   RUNG wire#powerrail
      Contact( "pH-2021_DB".Alarms.HighHigh )
   END_RUNG wire#w20
   RUNG wire#powerrail
      { S7_Templates := "SrcType := Time" } GE_Contact(in1 := "VFD-R201_DB".TIMEOUT.PT, in2 := T#8s)
   END_RUNG wire#w21
   RUNG wire#powerrail
      { S7_Templates := "SrcType := Time" } GE_Contact(in1 := "P-201A_DB".CF_Delay_TON.ET, in2 := T#8s)
   END_RUNG wire#w22
   RUNG wire#powerrail
      { S7_Templates := "SrcType := Time" } GE_Contact(in1 := "P-201B_DB".CF_Delay_TON.ET, in2 := T#8s)
   END_RUNG wire#w23
   RUNG wire#powerrail
      I_Contact( "T-101_Interlocks_DB".Out )
      P_Trig( "R-201_DB".OS.bit[1] )
   END_RUNG wire#w24
   // the same network as SCL:
   #_w1 := NOT "T-101_Interlocks_DB".Out AND NOT "R-201_DB".OS.bit[1];   // rising edge
   "R-201_DB".OS.bit[1] := NOT "T-101_Interlocks_DB".Out;
   "R-201_Interlocks_DB"(Interlock_1 := "LT-2011_DB".Alarms.HighHigh,   // "Interlocks"
                         Interlock_2 := "LSHH-2011_DB".Q,
                         Interlock_3 := "PT-201A_DB".Alarms.HighHigh,
                         Interlock_4 := "PT-201B_DB".Alarms.HighHigh,
                         Interlock_5 := "LT-2011_DB".Alarms.TransmitterFault,
                         Interlock_6 := "PT-201A_DB".Alarms.TransmitterFault,
                         Interlock_7 := "PT-201B_DB".Alarms.TransmitterFault,
                         Interlock_8 := "TT-2011_DB".Alarms.TransmitterFault,
                         Interlock_9 := "TT-2012_DB".Alarms.TransmitterFault,
                         Interlock_10 := "pH-2011_DB".Alarms.TransmitterFault,
                         Interlock_11 := "pH-2012_DB".Alarms.TransmitterFault,
                         Interlock_12 := "FT-2011_DB".Alarms.TransmitterFault,
                         Interlock_13 := "FT-2021_DB".Alarms.TransmitterFault,
                         Interlock_14 := "XV-2021_DB".Alarms."TO" OR "XV-2021_DB".Alarms.TC,
                         Interlock_15 := "XV-2013_DB".Alarms."TO" OR "XV-2013_DB".Alarms.TC,
                         Interlock_16 := "XV-1043_DB".Alarms."TO" OR "XV-1043_DB".Alarms.TC,
                         Interlock_17 := "XV-2011_DB".Alarms."TO" OR "XV-2011_DB".Alarms.TC,
                         Interlock_18 := "FT-1043_DB".Alarms.TransmitterFault,
                         Interlock_19 := "pH-2022_DB".Alarms.HighHigh,
                         Interlock_20 := "pH-2021_DB".Alarms.HighHigh,
                         Interlock_21 := "VFD-R201_DB".TIMEOUT.PT >= T#8s,
                         Interlock_22 := "P-201A_DB".CF_Delay_TON.ET >= T#8s,
                         Interlock_23 := "P-201B_DB".CF_Delay_TON.ET >= T#8s,
                         Interlock_25 := #_w1);
END_REGION

REGION Network 2: R-202 as Unit Interlocks
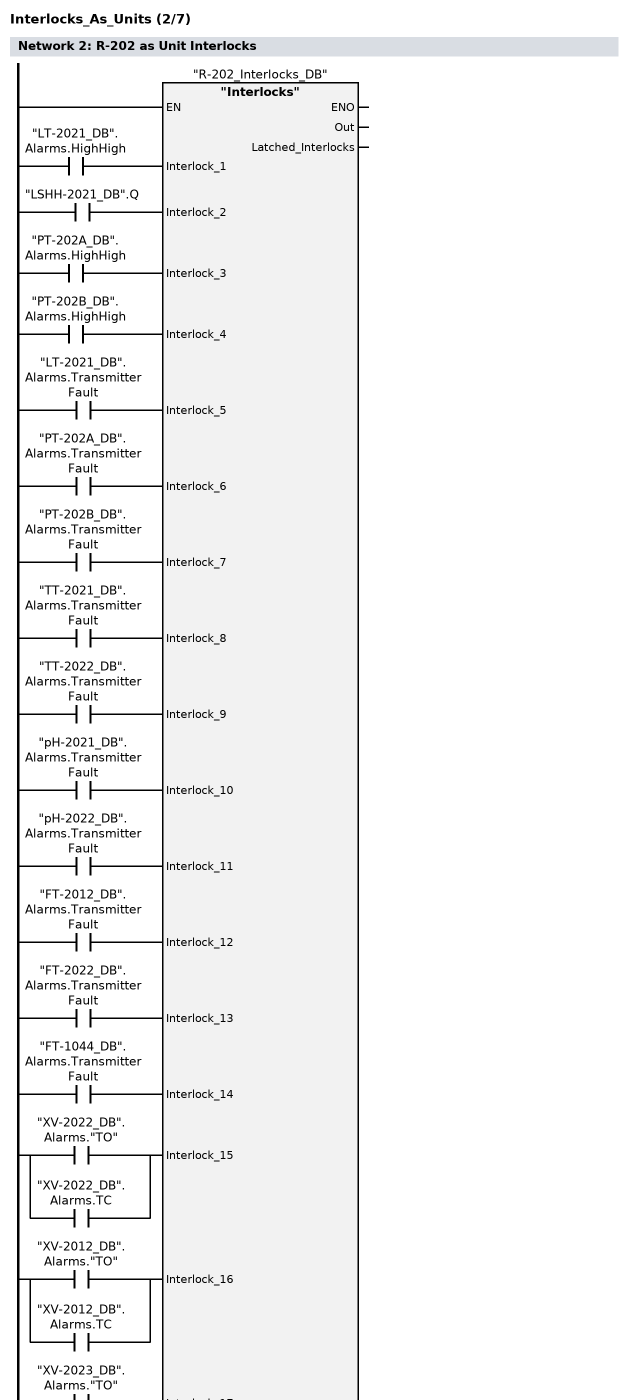
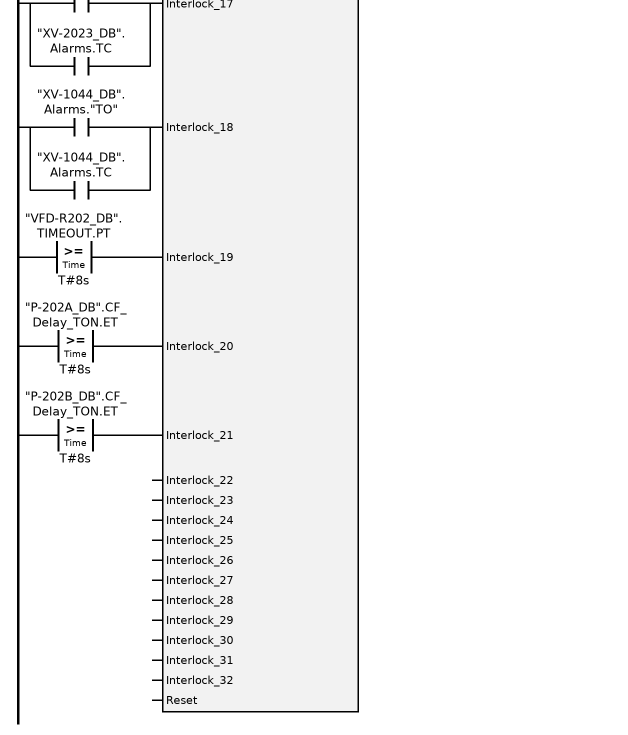
   RUNG wire#powerrail
      "R-202_Interlocks_DB"(Interlock_1 := wire#w1, Interlock_2 := wire#w2, Interlock_3 := wire#w3, Interlock_4 := wire#w4, Interlock_5 := wire#w5, Interlock_6 := wire#w6, Interlock_7 := wire#w7, Interlock_8 := wire#w8, Interlock_9 := wire#w9, Interlock_10 := wire#w10, Interlock_11 := wire#w11, Interlock_12 := wire#w12, Interlock_13 := wire#w13, Interlock_14 := wire#w14, Interlock_15 := wire#w15, Interlock_16 := wire#w16, Interlock_17 := wire#w17, Interlock_18 := wire#w18, Interlock_19 := wire#w19, Interlock_20 := wire#w20, Interlock_21 := wire#w21, Interlock_22 :=, Interlock_23 :=, Interlock_24 :=, Interlock_25 :=, Interlock_26 :=, Interlock_27 :=, Interlock_28 :=, Interlock_29 :=, Interlock_30 :=, Interlock_31 :=, Interlock_32 :=, Reset :=, Out =>, Latched_Interlocks =>)
   END_RUNG
   RUNG wire#powerrail
      Contact( "LT-2021_DB".Alarms.HighHigh )
   END_RUNG wire#w1
   RUNG wire#powerrail
      Contact( "LSHH-2021_DB".Q )
   END_RUNG wire#w2
   RUNG wire#powerrail
      Contact( "PT-202A_DB".Alarms.HighHigh )
   END_RUNG wire#w3
   RUNG wire#powerrail
      Contact( "PT-202B_DB".Alarms.HighHigh )
   END_RUNG wire#w4
   RUNG wire#powerrail
      Contact( "LT-2021_DB".Alarms.TransmitterFault )
   END_RUNG wire#w5
   RUNG wire#powerrail
      Contact( "PT-202A_DB".Alarms.TransmitterFault )
   END_RUNG wire#w6
   RUNG wire#powerrail
      Contact( "PT-202B_DB".Alarms.TransmitterFault )
   END_RUNG wire#w7
   RUNG wire#powerrail
      Contact( "TT-2021_DB".Alarms.TransmitterFault )
   END_RUNG wire#w8
   RUNG wire#powerrail
      Contact( "TT-2022_DB".Alarms.TransmitterFault )
   END_RUNG wire#w9
   RUNG wire#powerrail
      Contact( "pH-2021_DB".Alarms.TransmitterFault )
   END_RUNG wire#w10
   RUNG wire#powerrail
      Contact( "pH-2022_DB".Alarms.TransmitterFault )
   END_RUNG wire#w11
   RUNG wire#powerrail
      Contact( "FT-2012_DB".Alarms.TransmitterFault )
   END_RUNG wire#w12
   RUNG wire#powerrail
      Contact( "FT-2022_DB".Alarms.TransmitterFault )
   END_RUNG wire#w13
   RUNG wire#powerrail
      Contact( "FT-1044_DB".Alarms.TransmitterFault )
   END_RUNG wire#w14
   RUNG wire#powerrail
      Contact( "XV-2022_DB".Alarms."TO" )
   END_RUNG wire#w15
   RUNG wire#powerrail
      Contact( "XV-2022_DB".Alarms.TC )
   END_RUNG wire#w15
   RUNG wire#powerrail
      Contact( "XV-2012_DB".Alarms."TO" )
   END_RUNG wire#w16
   RUNG wire#powerrail
      Contact( "XV-2012_DB".Alarms.TC )
   END_RUNG wire#w16
   RUNG wire#powerrail
      Contact( "XV-2023_DB".Alarms."TO" )
   END_RUNG wire#w17
   RUNG wire#powerrail
      Contact( "XV-2023_DB".Alarms.TC )
   END_RUNG wire#w17
   RUNG wire#powerrail
      Contact( "XV-1044_DB".Alarms."TO" )
   END_RUNG wire#w18
   RUNG wire#powerrail
      Contact( "XV-1044_DB".Alarms.TC )
   END_RUNG wire#w18
   RUNG wire#powerrail
      { S7_Templates := "SrcType := Time" } GE_Contact(in1 := "VFD-R202_DB".TIMEOUT.PT, in2 := T#8s)
   END_RUNG wire#w19
   RUNG wire#powerrail
      { S7_Templates := "SrcType := Time" } GE_Contact(in1 := "P-202A_DB".CF_Delay_TON.ET, in2 := T#8s)
   END_RUNG wire#w20
   RUNG wire#powerrail
      { S7_Templates := "SrcType := Time" } GE_Contact(in1 := "P-202B_DB".CF_Delay_TON.ET, in2 := T#8s)
   END_RUNG wire#w21
   // the same network as SCL:
   "R-202_Interlocks_DB"(Interlock_1 := "LT-2021_DB".Alarms.HighHigh,   // "Interlocks"
                         Interlock_2 := "LSHH-2021_DB".Q,
                         Interlock_3 := "PT-202A_DB".Alarms.HighHigh,
                         Interlock_4 := "PT-202B_DB".Alarms.HighHigh,
                         Interlock_5 := "LT-2021_DB".Alarms.TransmitterFault,
                         Interlock_6 := "PT-202A_DB".Alarms.TransmitterFault,
                         Interlock_7 := "PT-202B_DB".Alarms.TransmitterFault,
                         Interlock_8 := "TT-2021_DB".Alarms.TransmitterFault,
                         Interlock_9 := "TT-2022_DB".Alarms.TransmitterFault,
                         Interlock_10 := "pH-2021_DB".Alarms.TransmitterFault,
                         Interlock_11 := "pH-2022_DB".Alarms.TransmitterFault,
                         Interlock_12 := "FT-2012_DB".Alarms.TransmitterFault,
                         Interlock_13 := "FT-2022_DB".Alarms.TransmitterFault,
                         Interlock_14 := "FT-1044_DB".Alarms.TransmitterFault,
                         Interlock_15 := "XV-2022_DB".Alarms."TO" OR "XV-2022_DB".Alarms.TC,
                         Interlock_16 := "XV-2012_DB".Alarms."TO" OR "XV-2012_DB".Alarms.TC,
                         Interlock_17 := "XV-2023_DB".Alarms."TO" OR "XV-2023_DB".Alarms.TC,
                         Interlock_18 := "XV-1044_DB".Alarms."TO" OR "XV-1044_DB".Alarms.TC,
                         Interlock_19 := "VFD-R202_DB".TIMEOUT.PT >= T#8s,
                         Interlock_20 := "P-202A_DB".CF_Delay_TON.ET >= T#8s,
                         Interlock_21 := "P-202B_DB".CF_Delay_TON.ET >= T#8s);
END_REGION

REGION Network 3: T-101 as Unit Iterlocks
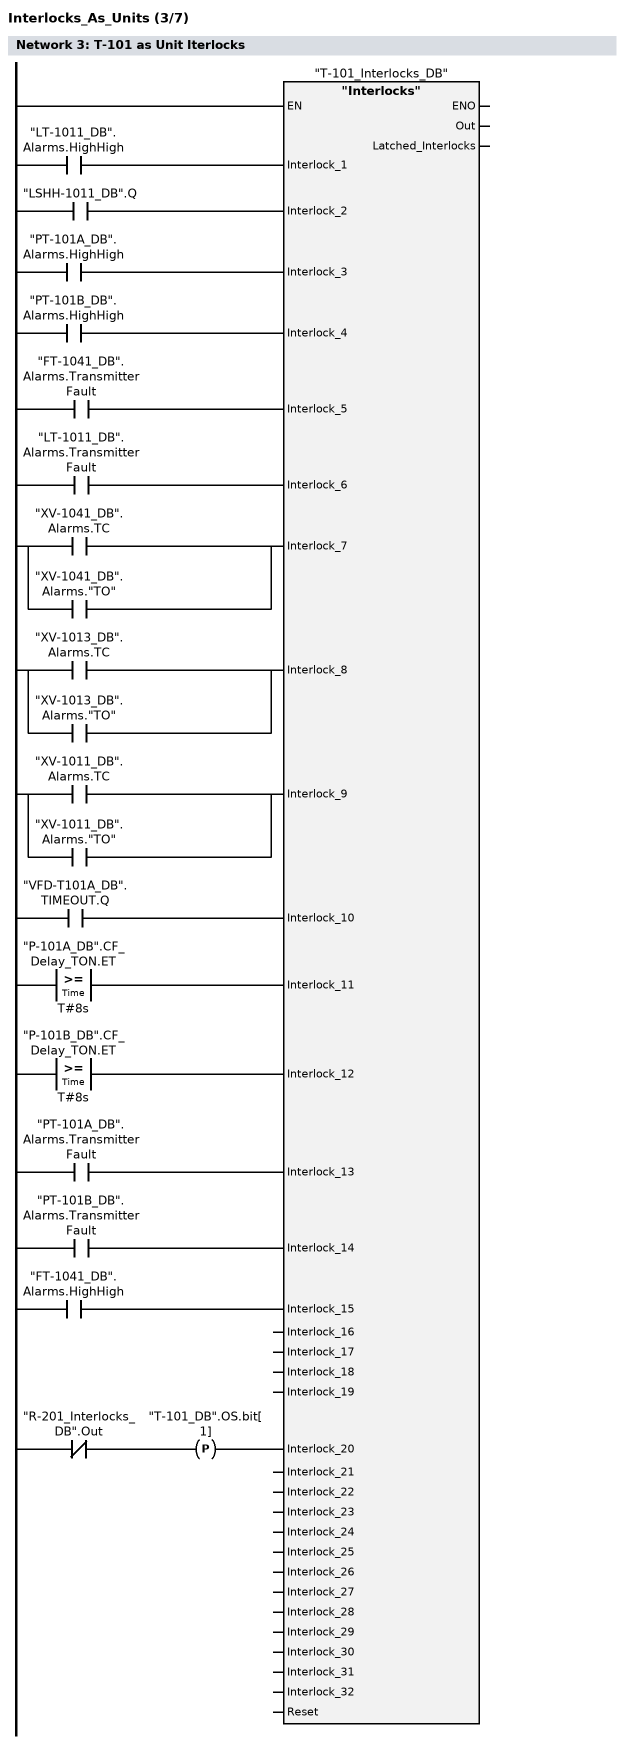
   RUNG wire#powerrail
      "T-101_Interlocks_DB"(Interlock_1 := wire#w1, Interlock_2 := wire#w2, Interlock_3 := wire#w3, Interlock_4 := wire#w4, Interlock_5 := wire#w5, Interlock_6 := wire#w6, Interlock_7 := wire#w7, Interlock_8 := wire#w8, Interlock_9 := wire#w9, Interlock_10 := wire#w10, Interlock_11 := wire#w11, Interlock_12 := wire#w12, Interlock_13 := wire#w13, Interlock_14 := wire#w14, Interlock_15 := wire#w15, Interlock_20 := wire#w16, Interlock_16 :=, Interlock_17 :=, Interlock_18 :=, Interlock_19 :=, Interlock_21 :=, Interlock_22 :=, Interlock_23 :=, Interlock_24 :=, Interlock_25 :=, Interlock_26 :=, Interlock_27 :=, Interlock_28 :=, Interlock_29 :=, Interlock_30 :=, Interlock_31 :=, Interlock_32 :=, Reset :=, Out =>, Latched_Interlocks =>)
   END_RUNG
   RUNG wire#powerrail
      Contact( "LT-1011_DB".Alarms.HighHigh )
   END_RUNG wire#w1
   RUNG wire#powerrail
      Contact( "LSHH-1011_DB".Q )
   END_RUNG wire#w2
   RUNG wire#powerrail
      Contact( "PT-101A_DB".Alarms.HighHigh )
   END_RUNG wire#w3
   RUNG wire#powerrail
      Contact( "PT-101B_DB".Alarms.HighHigh )
   END_RUNG wire#w4
   RUNG wire#powerrail
      Contact( "FT-1041_DB".Alarms.TransmitterFault )
   END_RUNG wire#w5
   RUNG wire#powerrail
      Contact( "LT-1011_DB".Alarms.TransmitterFault )
   END_RUNG wire#w6
   RUNG wire#powerrail
      Contact( "XV-1041_DB".Alarms.TC )
   END_RUNG wire#w7
   RUNG wire#powerrail
      Contact( "XV-1041_DB".Alarms."TO" )
   END_RUNG wire#w7
   RUNG wire#powerrail
      Contact( "XV-1013_DB".Alarms.TC )
   END_RUNG wire#w8
   RUNG wire#powerrail
      Contact( "XV-1013_DB".Alarms."TO" )
   END_RUNG wire#w8
   RUNG wire#powerrail
      Contact( "XV-1011_DB".Alarms.TC )
   END_RUNG wire#w9
   RUNG wire#powerrail
      Contact( "XV-1011_DB".Alarms."TO" )
   END_RUNG wire#w9
   RUNG wire#powerrail
      Contact( "VFD-T101A_DB".TIMEOUT.Q )
   END_RUNG wire#w10
   RUNG wire#powerrail
      { S7_Templates := "SrcType := Time" } GE_Contact(in1 := "P-101A_DB".CF_Delay_TON.ET, in2 := T#8s)
   END_RUNG wire#w11
   RUNG wire#powerrail
      { S7_Templates := "SrcType := Time" } GE_Contact(in1 := "P-101B_DB".CF_Delay_TON.ET, in2 := T#8s)
   END_RUNG wire#w12
   RUNG wire#powerrail
      Contact( "PT-101A_DB".Alarms.TransmitterFault )
   END_RUNG wire#w13
   RUNG wire#powerrail
      Contact( "PT-101B_DB".Alarms.TransmitterFault )
   END_RUNG wire#w14
   RUNG wire#powerrail
      Contact( "FT-1041_DB".Alarms.HighHigh )
   END_RUNG wire#w15
   RUNG wire#powerrail
      I_Contact( "R-201_Interlocks_DB".Out )
      P_Trig( "T-101_DB".OS.bit[1] )
   END_RUNG wire#w16
   // the same network as SCL:
   #_w1 := NOT "R-201_Interlocks_DB".Out AND NOT "T-101_DB".OS.bit[1];   // rising edge
   "T-101_DB".OS.bit[1] := NOT "R-201_Interlocks_DB".Out;
   "T-101_Interlocks_DB"(Interlock_1 := "LT-1011_DB".Alarms.HighHigh,   // "Interlocks"
                         Interlock_2 := "LSHH-1011_DB".Q,
                         Interlock_3 := "PT-101A_DB".Alarms.HighHigh,
                         Interlock_4 := "PT-101B_DB".Alarms.HighHigh,
                         Interlock_5 := "FT-1041_DB".Alarms.TransmitterFault,
                         Interlock_6 := "LT-1011_DB".Alarms.TransmitterFault,
                         Interlock_7 := "XV-1041_DB".Alarms.TC OR "XV-1041_DB".Alarms."TO",
                         Interlock_8 := "XV-1013_DB".Alarms.TC OR "XV-1013_DB".Alarms."TO",
                         Interlock_9 := "XV-1011_DB".Alarms.TC OR "XV-1011_DB".Alarms."TO",
                         Interlock_10 := "VFD-T101A_DB".TIMEOUT.Q,
                         Interlock_11 := "P-101A_DB".CF_Delay_TON.ET >= T#8s,
                         Interlock_12 := "P-101B_DB".CF_Delay_TON.ET >= T#8s,
                         Interlock_13 := "PT-101A_DB".Alarms.TransmitterFault,
                         Interlock_14 := "PT-101B_DB".Alarms.TransmitterFault,
                         Interlock_15 := "FT-1041_DB".Alarms.HighHigh,
                         Interlock_20 := #_w1);
END_REGION

REGION Network 4: T-102 as Unit Iterlocks
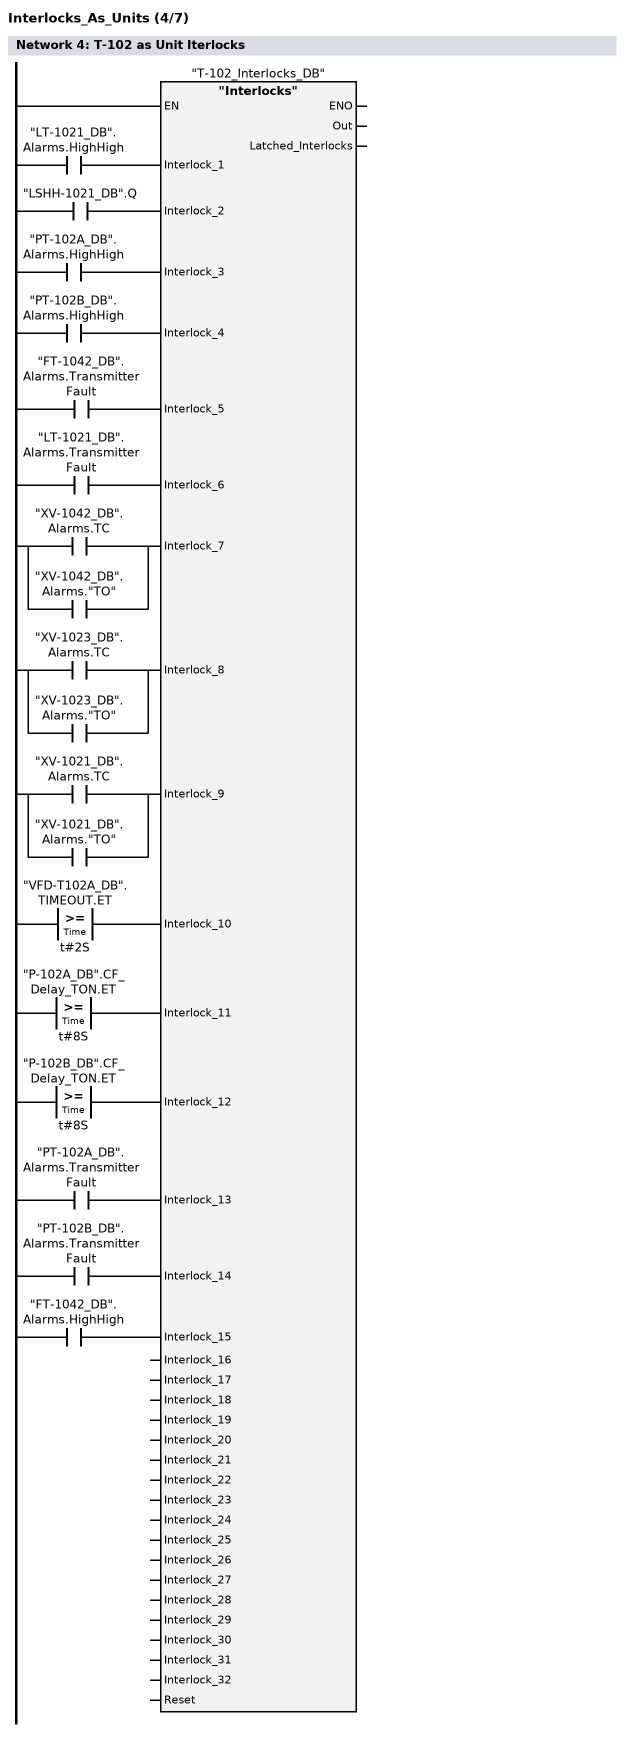
   RUNG wire#powerrail
      "T-102_Interlocks_DB"(Interlock_1 := wire#w1, Interlock_2 := wire#w2, Interlock_3 := wire#w3, Interlock_4 := wire#w4, Interlock_5 := wire#w5, Interlock_6 := wire#w6, Interlock_7 := wire#w7, Interlock_8 := wire#w8, Interlock_9 := wire#w9, Interlock_10 := wire#w10, Interlock_11 := wire#w11, Interlock_12 := wire#w12, Interlock_13 := wire#w13, Interlock_14 := wire#w14, Interlock_15 := wire#w15, Interlock_16 :=, Interlock_17 :=, Interlock_18 :=, Interlock_19 :=, Interlock_20 :=, Interlock_21 :=, Interlock_22 :=, Interlock_23 :=, Interlock_24 :=, Interlock_25 :=, Interlock_26 :=, Interlock_27 :=, Interlock_28 :=, Interlock_29 :=, Interlock_30 :=, Interlock_31 :=, Interlock_32 :=, Reset :=, Out =>, Latched_Interlocks =>)
   END_RUNG
   RUNG wire#powerrail
      Contact( "LT-1021_DB".Alarms.HighHigh )
   END_RUNG wire#w1
   RUNG wire#powerrail
      Contact( "LSHH-1021_DB".Q )
   END_RUNG wire#w2
   RUNG wire#powerrail
      Contact( "PT-102A_DB".Alarms.HighHigh )
   END_RUNG wire#w3
   RUNG wire#powerrail
      Contact( "PT-102B_DB".Alarms.HighHigh )
   END_RUNG wire#w4
   RUNG wire#powerrail
      Contact( "FT-1042_DB".Alarms.TransmitterFault )
   END_RUNG wire#w5
   RUNG wire#powerrail
      Contact( "LT-1021_DB".Alarms.TransmitterFault )
   END_RUNG wire#w6
   RUNG wire#powerrail
      Contact( "XV-1042_DB".Alarms.TC )
   END_RUNG wire#w7
   RUNG wire#powerrail
      Contact( "XV-1042_DB".Alarms."TO" )
   END_RUNG wire#w7
   RUNG wire#powerrail
      Contact( "XV-1023_DB".Alarms.TC )
   END_RUNG wire#w8
   RUNG wire#powerrail
      Contact( "XV-1023_DB".Alarms."TO" )
   END_RUNG wire#w8
   RUNG wire#powerrail
      Contact( "XV-1021_DB".Alarms.TC )
   END_RUNG wire#w9
   RUNG wire#powerrail
      Contact( "XV-1021_DB".Alarms."TO" )
   END_RUNG wire#w9
   RUNG wire#powerrail
      { S7_Templates := "SrcType := Time" } GE_Contact(in1 := "VFD-T102A_DB".TIMEOUT.ET, in2 := t#2S)
   END_RUNG wire#w10
   RUNG wire#powerrail
      { S7_Templates := "SrcType := Time" } GE_Contact(in1 := "P-102A_DB".CF_Delay_TON.ET, in2 := t#8S)
   END_RUNG wire#w11
   RUNG wire#powerrail
      { S7_Templates := "SrcType := Time" } GE_Contact(in1 := "P-102B_DB".CF_Delay_TON.ET, in2 := t#8S)
   END_RUNG wire#w12
   RUNG wire#powerrail
      Contact( "PT-102A_DB".Alarms.TransmitterFault )
   END_RUNG wire#w13
   RUNG wire#powerrail
      Contact( "PT-102B_DB".Alarms.TransmitterFault )
   END_RUNG wire#w14
   RUNG wire#powerrail
      Contact( "FT-1042_DB".Alarms.HighHigh )
   END_RUNG wire#w15
   // the same network as SCL:
   "T-102_Interlocks_DB"(Interlock_1 := "LT-1021_DB".Alarms.HighHigh,   // "Interlocks"
                         Interlock_2 := "LSHH-1021_DB".Q,
                         Interlock_3 := "PT-102A_DB".Alarms.HighHigh,
                         Interlock_4 := "PT-102B_DB".Alarms.HighHigh,
                         Interlock_5 := "FT-1042_DB".Alarms.TransmitterFault,
                         Interlock_6 := "LT-1021_DB".Alarms.TransmitterFault,
                         Interlock_7 := "XV-1042_DB".Alarms.TC OR "XV-1042_DB".Alarms."TO",
                         Interlock_8 := "XV-1023_DB".Alarms.TC OR "XV-1023_DB".Alarms."TO",
                         Interlock_9 := "XV-1021_DB".Alarms.TC OR "XV-1021_DB".Alarms."TO",
                         Interlock_10 := "VFD-T102A_DB".TIMEOUT.ET >= t#2S,
                         Interlock_11 := "P-102A_DB".CF_Delay_TON.ET >= t#8S,
                         Interlock_12 := "P-102B_DB".CF_Delay_TON.ET >= t#8S,
                         Interlock_13 := "PT-102A_DB".Alarms.TransmitterFault,
                         Interlock_14 := "PT-102B_DB".Alarms.TransmitterFault,
                         Interlock_15 := "FT-1042_DB".Alarms.HighHigh);
END_REGION

REGION Network 5: T-103 as Unit Iterlocks
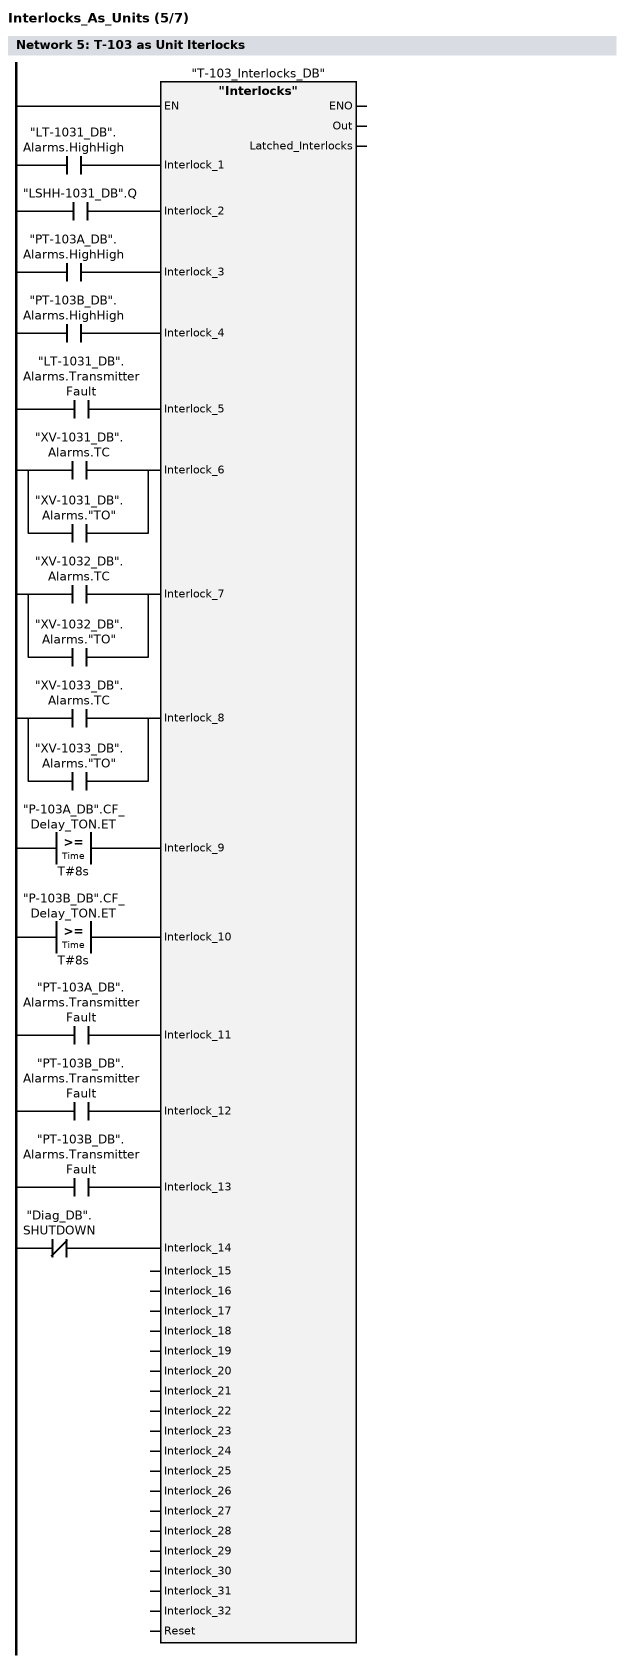
   RUNG wire#powerrail
      "T-103_Interlocks_DB"(Interlock_1 := wire#w1, Interlock_2 := wire#w2, Interlock_3 := wire#w3, Interlock_4 := wire#w4, Interlock_5 := wire#w5, Interlock_6 := wire#w6, Interlock_7 := wire#w7, Interlock_8 := wire#w8, Interlock_9 := wire#w9, Interlock_10 := wire#w10, Interlock_11 := wire#w11, Interlock_12 := wire#w12, Interlock_13 := wire#w13, Interlock_14 := wire#w14, Interlock_15 :=, Interlock_16 :=, Interlock_17 :=, Interlock_18 :=, Interlock_19 :=, Interlock_20 :=, Interlock_21 :=, Interlock_22 :=, Interlock_23 :=, Interlock_24 :=, Interlock_25 :=, Interlock_26 :=, Interlock_27 :=, Interlock_28 :=, Interlock_29 :=, Interlock_30 :=, Interlock_31 :=, Interlock_32 :=, Reset :=, Out =>, Latched_Interlocks =>)
   END_RUNG
   RUNG wire#powerrail
      Contact( "LT-1031_DB".Alarms.HighHigh )
   END_RUNG wire#w1
   RUNG wire#powerrail
      Contact( "LSHH-1031_DB".Q )
   END_RUNG wire#w2
   RUNG wire#powerrail
      Contact( "PT-103A_DB".Alarms.HighHigh )
   END_RUNG wire#w3
   RUNG wire#powerrail
      Contact( "PT-103B_DB".Alarms.HighHigh )
   END_RUNG wire#w4
   RUNG wire#powerrail
      Contact( "LT-1031_DB".Alarms.TransmitterFault )
   END_RUNG wire#w5
   RUNG wire#powerrail
      Contact( "XV-1031_DB".Alarms.TC )
   END_RUNG wire#w6
   RUNG wire#powerrail
      Contact( "XV-1031_DB".Alarms."TO" )
   END_RUNG wire#w6
   RUNG wire#powerrail
      Contact( "XV-1032_DB".Alarms.TC )
   END_RUNG wire#w7
   RUNG wire#powerrail
      Contact( "XV-1032_DB".Alarms."TO" )
   END_RUNG wire#w7
   RUNG wire#powerrail
      Contact( "XV-1033_DB".Alarms.TC )
   END_RUNG wire#w8
   RUNG wire#powerrail
      Contact( "XV-1033_DB".Alarms."TO" )
   END_RUNG wire#w8
   RUNG wire#powerrail
      { S7_Templates := "SrcType := Time" } GE_Contact(in1 := "P-103A_DB".CF_Delay_TON.ET, in2 := T#8s)
   END_RUNG wire#w9
   RUNG wire#powerrail
      { S7_Templates := "SrcType := Time" } GE_Contact(in1 := "P-103B_DB".CF_Delay_TON.ET, in2 := T#8s)
   END_RUNG wire#w10
   RUNG wire#powerrail
      Contact( "PT-103A_DB".Alarms.TransmitterFault )
   END_RUNG wire#w11
   RUNG wire#powerrail
      Contact( "PT-103B_DB".Alarms.TransmitterFault )
   END_RUNG wire#w12
   RUNG wire#powerrail
      Contact( "PT-103B_DB".Alarms.TransmitterFault )
   END_RUNG wire#w13
   RUNG wire#powerrail
      I_Contact( "Diag_DB".SHUTDOWN )
   END_RUNG wire#w14
   // the same network as SCL:
   "T-103_Interlocks_DB"(Interlock_1 := "LT-1031_DB".Alarms.HighHigh,   // "Interlocks"
                         Interlock_2 := "LSHH-1031_DB".Q,
                         Interlock_3 := "PT-103A_DB".Alarms.HighHigh,
                         Interlock_4 := "PT-103B_DB".Alarms.HighHigh,
                         Interlock_5 := "LT-1031_DB".Alarms.TransmitterFault,
                         Interlock_6 := "XV-1031_DB".Alarms.TC OR "XV-1031_DB".Alarms."TO",
                         Interlock_7 := "XV-1032_DB".Alarms.TC OR "XV-1032_DB".Alarms."TO",
                         Interlock_8 := "XV-1033_DB".Alarms.TC OR "XV-1033_DB".Alarms."TO",
                         Interlock_9 := "P-103A_DB".CF_Delay_TON.ET >= T#8s,
                         Interlock_10 := "P-103B_DB".CF_Delay_TON.ET >= T#8s,
                         Interlock_11 := "PT-103A_DB".Alarms.TransmitterFault,
                         Interlock_12 := "PT-103B_DB".Alarms.TransmitterFault,
                         Interlock_13 := "PT-103B_DB".Alarms.TransmitterFault,
                         Interlock_14 := NOT "Diag_DB".SHUTDOWN);
END_REGION

REGION Network 6: T-104 as Unit Iterlocks
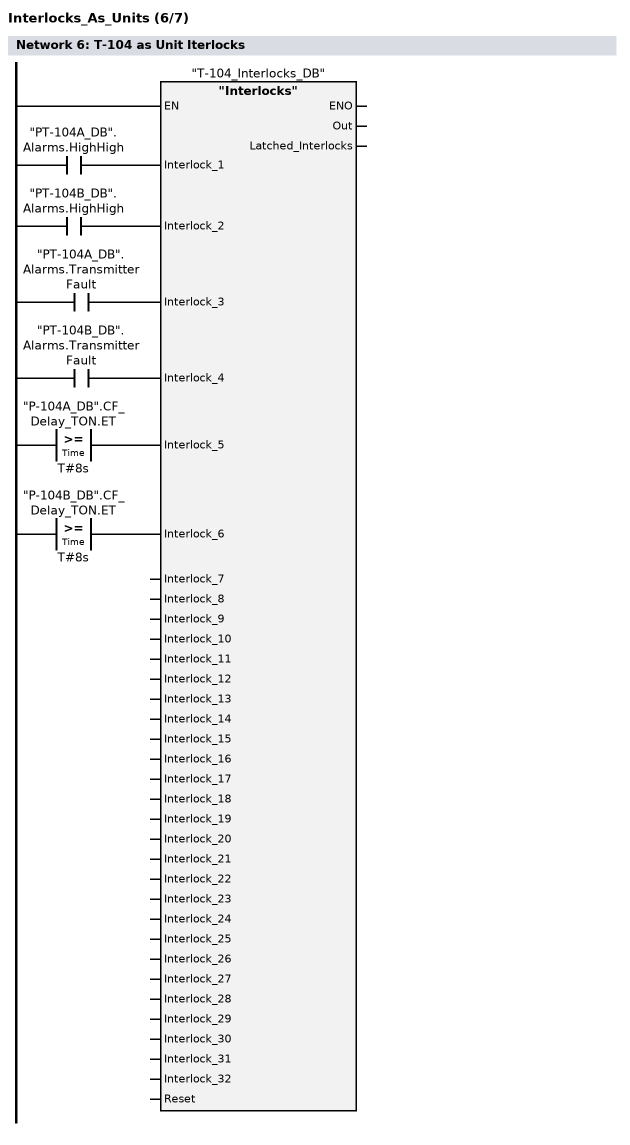
   RUNG wire#powerrail
      "T-104_Interlocks_DB"(Interlock_1 := wire#w1, Interlock_2 := wire#w2, Interlock_3 := wire#w3, Interlock_4 := wire#w4, Interlock_5 := wire#w5, Interlock_6 := wire#w6, Interlock_7 :=, Interlock_8 :=, Interlock_9 :=, Interlock_10 :=, Interlock_11 :=, Interlock_12 :=, Interlock_13 :=, Interlock_14 :=, Interlock_15 :=, Interlock_16 :=, Interlock_17 :=, Interlock_18 :=, Interlock_19 :=, Interlock_20 :=, Interlock_21 :=, Interlock_22 :=, Interlock_23 :=, Interlock_24 :=, Interlock_25 :=, Interlock_26 :=, Interlock_27 :=, Interlock_28 :=, Interlock_29 :=, Interlock_30 :=, Interlock_31 :=, Interlock_32 :=, Reset :=, Out =>, Latched_Interlocks =>)
   END_RUNG
   RUNG wire#powerrail
      Contact( "PT-104A_DB".Alarms.HighHigh )
   END_RUNG wire#w1
   RUNG wire#powerrail
      Contact( "PT-104B_DB".Alarms.HighHigh )
   END_RUNG wire#w2
   RUNG wire#powerrail
      Contact( "PT-104A_DB".Alarms.TransmitterFault )
   END_RUNG wire#w3
   RUNG wire#powerrail
      Contact( "PT-104B_DB".Alarms.TransmitterFault )
   END_RUNG wire#w4
   RUNG wire#powerrail
      { S7_Templates := "SrcType := Time" } GE_Contact(in1 := "P-104A_DB".CF_Delay_TON.ET, in2 := T#8s)
   END_RUNG wire#w5
   RUNG wire#powerrail
      { S7_Templates := "SrcType := Time" } GE_Contact(in1 := "P-104B_DB".CF_Delay_TON.ET, in2 := T#8s)
   END_RUNG wire#w6
   // the same network as SCL:
   "T-104_Interlocks_DB"(Interlock_1 := "PT-104A_DB".Alarms.HighHigh,   // "Interlocks"
                         Interlock_2 := "PT-104B_DB".Alarms.HighHigh,
                         Interlock_3 := "PT-104A_DB".Alarms.TransmitterFault,
                         Interlock_4 := "PT-104B_DB".Alarms.TransmitterFault,
                         Interlock_5 := "P-104A_DB".CF_Delay_TON.ET >= T#8s,
                         Interlock_6 := "P-104B_DB".CF_Delay_TON.ET >= T#8s);
END_REGION

REGION Network 7: Centrifuge Interlocks
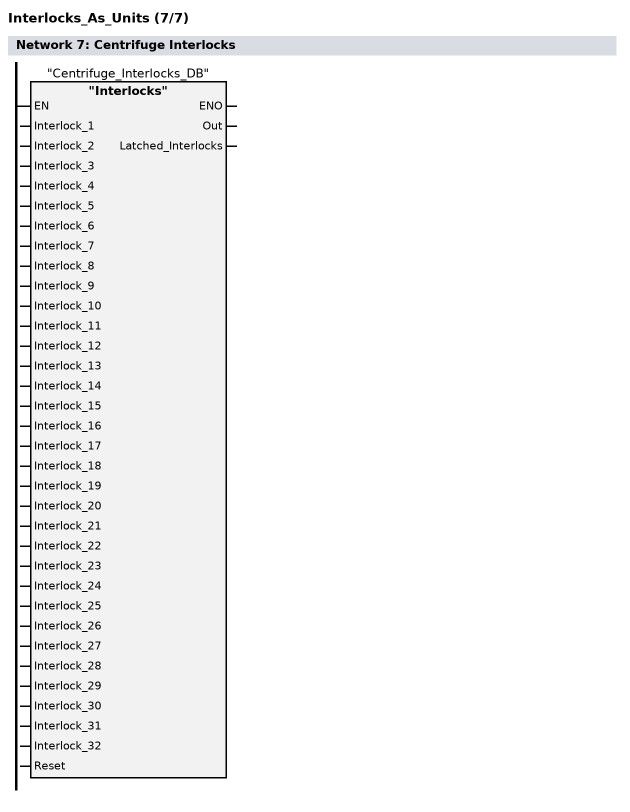
   RUNG wire#powerrail
      "Centrifuge_Interlocks_DB"(Interlock_1 :=, Interlock_2 :=, Interlock_3 :=, Interlock_4 :=, Interlock_5 :=, Interlock_6 :=, Interlock_7 :=, Interlock_8 :=, Interlock_9 :=, Interlock_10 :=, Interlock_11 :=, Interlock_12 :=, Interlock_13 :=, Interlock_14 :=, Interlock_15 :=, Interlock_16 :=, Interlock_17 :=, Interlock_18 :=, Interlock_19 :=, Interlock_20 :=, Interlock_21 :=, Interlock_22 :=, Interlock_23 :=, Interlock_24 :=, Interlock_25 :=, Interlock_26 :=, Interlock_27 :=, Interlock_28 :=, Interlock_29 :=, Interlock_30 :=, Interlock_31 :=, Interlock_32 :=, Reset :=, Out =>, Latched_Interlocks =>)
   END_RUNG
   // the same network as SCL:
   "Centrifuge_Interlocks_DB"();   // "Interlocks"
END_REGION

REGION Network 8 (SCL): Units Interlocks
   //Interlocks to the Units
   //T-101
   "T-101_DB".Cmds.IL := "T-101 Mix & Wash X material INTERLOCKS".Out AND "T-101_DB".Cmds.PermCond;
   //T-102
   "T-102_DB".Cmds.IL := "T-102 Mix & Wash Y Material  INTERLOCKS".Out AND "T-102_DB".Cmds.PermCond;
   //T-103
   "T-103_DB".Cmds.IL:= "T-103_Interlocks_DB".Out AND "T-103_DB".Cmds.PermCond;
   //T-104
   "T-104_DB".Cmds.IL := "T-104_Interlocks_DB".Out AND "T-104_DB".Cmds.PermCond;
   //R-201
   "R-201_DB".Cmds.IL := "I201A_Reactor_Interlocks".Out AND "I201B_Reactor_Interlocks".Out AND "R-201_DB".Cmds.PermCond;
   //R-202
   "R-202_DB".Cmds.IL := "I202A_Reactors_Interlocks".Out AND "I202B_Reactors_Interlocks".Out AND "R-202_DB".Cmds.PermCond;
   //Centrifuge
   "Centrifuge_DB".Cmds.IL := "C-301 Centrifuge_INTERLOCKS".Out AND "Centrifuge_DB".Cmds.PermCond;
   //R-401
   "R-401_DB".Cmds.IL :=  "I401_Calcination_Interlocks".Out AND "R-401_DB".Cmds.PermCond;
   //R-402
   "R-402_DB".Cmds.IL := "I402_Passivate_Interlocks".Out AND "R-402_DB".Cmds.PermCond;
END_REGION
END_FUNCTION

// folder: Outside Comms/Centrifuge

FUNCTION "ExchangeCentrifuge_FC" : Void   // FC34, LAD
{ S7_Optimized_Access := 'TRUE' }
VERSION : 0.1
   VAR_TEMP
      ss : Bool;
      estp : Bool;
      reset : Bool;
      fe : Bool;
      sp : Int;
      FromC : Struct
         vf : Bool;
         estop : Bool;
         sfault : Bool;
         bskf : Bool;
         conl : Bool;
         fr : Bool;
         vt : Int;
         pv : Int;
      END_STRUCT;
   END_VAR
BEGIN

REGION Network 2: ////*********From DCS to Centrifuge**********////
   // Periphery Signal will be added to the coils.
END_REGION

REGION Network 3: Start/Stop Command